   63: 'El compresor Sullair 1 superó la máxima cantidad de horas sin mantenimiento #1', class MTA, trigger "Rec21" bit 13
   64: 'El compresor Sullair 1 superó la máxima cantidad de horas sin mantenimiento #2', class MTA, trigger "Rec21" bit 14
   65: 'El compresor Sullair 1 superó la máxima cantidad de horas sin mantenimiento #3', class MTA, trigger "Rec21" bit 15
   84: 'El compresor Sullair 1 superó la máxima cantidad de horas sin mantenimiento #4', class MTA, trigger "Rec22" bit 8
   85: 'El compresor Sullair 1 superó la máxima cantidad de horas sin mantenimiento #5', class MTA, trigger "Rec22" bit 9
   86: 'El compresor Sullair 0 superó la máxima cantidad de horas sin mantenimiento #1', class MTA, trigger "Rec22" bit 10
   122: 'El compresor Sullair 0 superó la máxima cantidad de horas sin mantenimiento #2', class MTA, trigger "Rec22" bit 11
   123: 'El compresor Sullair 0 superó la máxima cantidad de horas sin mantenimiento #3', class MTA, trigger "Rec22" bit 12
   124: 'El compresor Sullair 0 superó la máxima cantidad de horas sin mantenimiento #4', class MTA, trigger "Rec22" bit 13
   173: 'El compresor Sullair 0 superó la máxima cantidad de horas sin mantenimiento #5', class MTA, trigger "Rec22" bit 14
   174: 'El compresor Atlas 3 superó la máxima cantidad de horas sin mantenimiento #1', class MTA, trigger "Rec22" bit 15
   175: 'El compresor Atlas 3 superó la máxima cantidad de horas sin mantenimiento #2', class MTA, trigger "Rec23" bit 8
   176: 'El compresor Atlas 3 superó la máxima cantidad de horas sin mantenimiento #3', class MTA, trigger "Rec23" bit 9
   177: 'El compresor Atlas 3 superó la máxima cantidad de horas sin mantenimiento #4', class MTA, trigger "Rec23" bit 10
   178: 'El compresor Atlas 3 superó la máxima cantidad de horas sin mantenimiento #5', class MTA, trigger "Rec23" bit 11
   179: 'El compresor Atlas 2 superó la máxima cantidad de horas sin mantenimiento #1', class MTA, trigger "Rec23" bit 12
   180: 'El compresor Atlas 2 superó la máxima cantidad de horas sin mantenimiento #2', class MTA, trigger "Rec23" bit 13
   181: 'El compresor Atlas 2 superó la máxima cantidad de horas sin mantenimiento #3', class MTA, trigger "Rec23" bit 14
   182: 'El compresor Atlas 2 superó la máxima cantidad de horas sin mantenimiento #4', class MTA, trigger "Rec23" bit 15
   183: 'El compresor Atlas 2 superó la máxima cantidad de horas sin mantenimiento #5', class MTA, trigger "Rec24" bit 8
   184: 'El booster 1 superó la máxima cantidad de horas sin mantenimiento', class MTA, trigger "Rec24" bit 9
   185: 'El booster 2 superó la máxima cantidad de horas sin mantenimiento', class MTA, trigger "Rec24" bit 10
   186: 'Temperatura agua de torres compresores elevada', class MTA, trigger "Rec24" bit 11
   187: 'Falla Confirmación de purga - ABC2', class MTA, trigger "Rec17" bit 8
   188: 'Falla Confirmación de purga - ABC3', class MTA, trigger "Rec17" bit 9
   189: 'Falla Confirmación de purga - Bellis', class MTA, trigger "Rec17" bit 10
   190: 'Falla Confirmación de purga - ABC4', class MTA, trigger "Rec17" bit 11
   191: 'Falla Confirmación de purga - ABC5', class MTA, trigger "Rec17" bit 12
   192: 'Falla Confirmación de purga - ABC1', class MTA, trigger "Rec17" bit 13
   199: 'Falla por relé de freq. Comp ALTA', class MTA, trigger "Rec24" bit 15

text list "EstadoMotor": 0 'Detenido'; 1 'En Marcha'; 2 'Arrancando'; 3 'Deteniéndose'; 4 'Espera para Arrancar'; 5 'Sobrecarga de Corriente'; 6 'Deshabilitado'; 7 'En Falla'

text list "EstadoCmpAlta": 256 'Manual'; 512 'Sin Requerimiento'; 1024 'Sin Marcha'; 2048 'En Vacío'; 4096 'En Carga'; 8192 'Manual sin Requerimiento'; 16384 ''; 32768 'Falla'; 1 'Requiere Marcha'

text list "Presostato Ctrl": 0 'Presostato de Control: Desactivado'; 1 'Presostato de Control: Activado'

text list "Presostato de Alarma": 0 'Presostato de Presión Alta: Activado'; 1 'Presostato de Presión Alta: Desactivado'

text list "Lista de rutas": 0 '\Storage Card USB\ABC-1\'; 1 '\Storage Card USB\ABC-2\'; 2 '\Storage Card USB\ABC-3\'; 3 '\Storage Card USB\ABC-4\'; 4 '\Storage Card USB\ABC-5\'; 5 '\Storage Card USB\Bellis\'; 6 '\Storage Card USB\Atlas2\'; 7 '\Storage Card USB\Atlas3\'; 8 '\Storage Card USB\Sullair0\'; 9 '\Storage Card USB\Sullair1\'; 10 '\Storage Card USB\Sullair2\'

text list "Lista de compresores": 0 'ABC-1'; 1 'ABC-2'; 2 'ABC-3'; 3 'ABC-4'; 4 'ABC-5'; 5 'Bellis'; 6 'Atlas 2'; 7 'Atlas 3'; 8 'Sullair 0'; 9 'Sullair 1'; 10 'Sullair 2'

graphic list "Motor2": 0 'Motor2Dorado'; 1 'Motor2Verde_1'; 2 'Motor2VerdeOscuro'; 3 'Motor2Azul'; 4 'Motor2Celeste'; 5 'Motor2Amarillo'; 6 'Motor2Gris_1'; 7 'Motor2Rojo'; 8 'Motor2Dorado'

graphic list "MotorBelliss": 0 'dorado'; 1 'bell1ve'; 2 'bell1ve'; 3 'az'; 4 'az'; 5 'bell1am'; 6 'dorado'; 7 'az'

graphic list "BarraPrioridades": 1 'R1'; 2 'R2'; 3 'R3'; 4 'R4'; 5 'R5'; 6 'R4'; 6 'R6.rlu'

graphic list "Indicador": 0 'indDorado'; 1 'indVerde'; 2 'indVerde_1'; 3 'indAZUL'; 4 'indCeleste'; 5 'indAmarillo'; 6 'indGris'; 7 'indRojo'; 8 'indCeleste'

graphic list "BarraPrioridades_1": 1 'set1'; 2 'set2'; 3 'set3'; 4 'set4'; 5 'set5'; 6 'set4'; 6 'set6'

graphic list "BaseSullChico": 0 'BaseSullChicoDorado_4'; 1 'BaseSullChico'; 2 'BaseSullChico'; 3 'BaseSullChicoAzul_4'; 4 'BaseSullChicoAzul_4'; 5 'BaseSullChicoAmarillo_4'; 6 'BaseSullChicoGris_4'; 7 'BaseSullChicoRojo_4'; 8 'BaseSullChicoAzul_4'

graphic list "MotorTorre": 0 'torreFINAL4C2_1'; 1 'torreFINAL4C2v_2'; 2 'torreFINAL4C2v_2'; 3 'torreFINAL4C2b'; 4 'torreFINAL4C2b'; 5 'torreFINAL4C2a_2'; 6 'torreFINAL4C2_1'; 7 'torreFINAL4C2_1'

graphic list "Secador2": 0 'BaseSullChicoDorado_2'; 1 'BaseSullChico_5'; 2 'BaseSullChico_5'; 3 'BaseSullChicoAzul_2'; 4 'BaseSullChicoAzul_2'; 5 'BaseSullChicoAmarillo_2'; 6 'BaseSullChicoGris_2'; 7 'BaseSullChicoRojo_2'

graphic list "Secador1": 0 'BaseSullChicoDorado_1'; 1 'BaseSullChico_4'; 2 'BaseSullChico_4'; 3 'BaseSullChicoAzul_1'; 4 'BaseSullChicoAzul_1'; 5 'BaseSullChicoAmarillo_1'; 6 'BaseSullChicoGris_1'; 7 'BaseSullChicoRojo_1'

graphic list "Motor Grande": 0 'MotorDorado'; 1 'MotorVerde'; 2 'MotorVerde'; 3 'MotorAzul'; 4 'MotorCeleste'; 5 'MotorAmarillo'; 6 'MotorGris'; 7 'MotorRojo'; 8 'MotorCeleste'

graphic list "Mantenimiento": 0 'MECH2'; 1 'MECH1'

graphic list "Motor Chico": 0 'Booster-D-Dor2'; 1 'Booster-D-VE2'; 2 'Booster-D-VE2'; 3 'Booster-D-Azul2'; 4 'Booster-D-AZ2'; 5 'Booster-D-AM2'; 6 'Booster-D-GR'; 7 'Booster-D-RO2'; 8 'Booster-D-AZ2'

graphic list "Hélice": 0 'Booster-C1'; 1 'Booster-C2'

screen "Graf-Corrientes" 1280x800, template "Plantilla"
   TrendView "Visor de curvas_1" at 8,72 size 1260x636
   TextField "Campo de texto_16" at 493,10 size 294x27; Text 'Gráficas - Sentron Pac - Corrientes'

screen "Graf-Fase" 1280x800, template "Plantilla"
   TrendView "Visor de curvas_1" at 3,65 size 1268x644
   TextField "Campo de texto_16" at 477,10 size 364x27; Text 'Gráficas - Sentron Pac - Tensiones de Fase'

screen "Grafica" 1280x800, template "Plantilla"
   Button "Botón_7" at 368,280 size 240x49; TextOff 'Presión Baja'
      on Click: ActivateScreen("GraficaPBAJA", 0)
   Button "Botón_12" at 367,440 size 240x49; TextOff 'Temperatura Chillers'
      on Click: ActivateScreen("GraficaTCH", 0)
   Button "Botón_13" at 368,216 size 240x49; TextOff 'Presión Alta'
      on Click: ActivateScreen("GraficaPALTA", 0)
   TextField "Campo de texto_1" at 55,108 size 353x27; Text 'Seleccione la variable que desea graficar:'
   Button "Botón_1" at 767,280 size 240x49; TextOff 'Todas Cavaleto'
      on Click: ActivateScreen("GraficaTodas", 0)
   TextField "Campo de texto_16" at 521,10 size 226x27; Text 'Graficar variable analógica'
   Button "Botón_2" at 368,344 size 240x49; TextOff 'Temperatura Cavaleto'
      on Click: ActivateScreen("GraficaTCAV", 0)
   Button "Botón_3" at 766,440 size 240x49; TextOff 'Grafico Caudal/Potencia'
      on Click: ActivateScreen("Graf-cau-pot-actual", 0)
   Button "Botón_4" at 769,526 size 240x49; TextOff 'Historico Caudal/Potencia'
      on Click: ActivateScreen("Graf-cau-pot-historico", 0)

screen "GraficaPALTA" 1280x800, template "Plantilla"
   TrendView "Visor de curvas_1" at 5,79 size 1234x618
   TextField "Campo de texto_16" at 521,10 size 193x27; Text 'Grafica Presión de Alta'

screen "GraficaPBAJA" 1280x800, template "Plantilla"
   TrendView "Visor de curvas_1" at 5,71 size 1242x626
   TextField "Campo de texto_16" at 521,10 size 198x27; Text 'Grafica Presión de Baja'

screen "GraficaTCAV" 1280x800, template "Plantilla"
   TrendView "Visor de curvas_1" at 5,71 size 1242x626
   TextField "Campo de texto_16" at 521,10 size 254x27; Text 'Grafica Temperatura Cavaleto'

screen "GraficaTCH" 1280x800, template "Plantilla"
   TrendView "Visor de curvas_1" at 5,71 size 1242x626
   TextField "Campo de texto_16" at 521,10 size 243x27; Text 'Grafica Temperatura Chillers'

screen "GraficaTodas" 1280x800, template "Plantilla"
   TrendView "Visor de curvas_1" at 5,71 size 1242x626

screen "Graf-Linea" 1280x800, template "Plantilla"
   TrendView "Visor de curvas_1" at 3,65 size 1268x652
   TextField "Campo de texto_16" at 453,10 size 370x27; Text 'Gráficas - Sentron Pac - Tensiones de Línea'

screen "Graf-Pot" 1280x800, template "Plantilla"
   TrendView "Visor de curvas_1" at 3,65 size 1268x644
   TextField "Campo de texto_16" at 477,10 size 339x27; Text 'Gráficas - Sentron Pac - Potencia x Fase'

screen "Graf-PotTotal" 1280x800, template "Plantilla"
   TrendView "Visor de curvas_1" at 3,65 size 1268x644
   TextField "Campo de texto_16" at 477,10 size 327x27; Text 'Gráficas - Sentron Pac - Potencia Total'

screen "IluminaciónMTA" 1280x800, template "Plantilla"
   Polygon "Polígono_6" at 1018,121 size 183x209
      Visibility <- "ON"
   Ellipse "Elipse_4" at 1019,317 size 184x29
      Visibility <- "ON"
   Polygon "Polígono_3" at 782,137 size 351x377
      Visibility <- "ON"
   Ellipse "Elipse_5" at 789,485 size 344x61
      Visibility <- "ON"
   Polygon "Polígono_2" at 446,161 size 559x577
      Visibility <- "ON"
   Ellipse "Elipse_1" at 694,118 size 59x74
      Appearance <- "ON"
   Ellipse "Elipse_2" at 940,112 size 35x50
      Appearance <- "ON"
   Ellipse "Elipse_3" at 1100,112 size 19x26
      Appearance <- "ON"
   Switch "Interruptor_1" at 36,546 size 510x96; TextOff 'Encendido Permanente OFF'; CaptionText 'Switch'; TextOn 'Encendido Permanente ON'
      Appearance <- "MantenerON"
      ProcessValue <- "MantenerON"
   Button "Botón_1" at 36,264 size 248x96; TextOff 'Encender'
      on Press: SetBit("EncendidoPanel")
      on Release: ResetBit("EncendidoPanel")
   Button "Botón_2" at 298,263 size 248x96; TextOff 'Apagar'
      on Press: SetBit("ApagadoPanel")
      on Release: ResetBit("ApagadoPanel")
   IOField "Campo ES_1" at 257,148 size 140x39; FormatPattern 99; Unit    Min.
      ProcessValue <- "TiempoIluminación"
   TextField "Campo de texto_1" at 42,156 size 186x27; Text 'Tiempo de encendido'
   TextField "Campo de texto_3" at 58,190 size 466x58; Text 'La iluminación puede ser encendida desde el panel o desde el pulsador. En caso de no ser apagada mediante los mismos medios, el PLC la apagará automáticamente al concluir el "tiempo de encendido".'
   TextField "Campo de texto_2" at 58,414 size 433x112; Text 'En caso de necesitar permanecer con la iluminación encendida durante un tiempo mayor al "tiempo de encendido", se provee la posibilidad de seleccionar el "encendido permanente". Mientras el "encendido permanente" esté activado la iluminación se mantendrá encendida, y el PLC dejará de controlar el apagado automático.'
   TextField "Campo de texto_16" at 553,10 size 177x27; Text 'Iluminación Cavaleto'

screen "INICIO" 1280x800, template "Plantilla"
   Button "Botón_1" at 1025,513 size 108x65; TextOff 'Cerrar Runtime'; Authorization "Administración de usuarios"
      on Press: StopRuntime(0)
   Button "Botón_2" at 115,501 size 130x47; TextOff 'Iniciar Sesion'; PictureOff "Gráfico_5"
      on Click: function_a2a04561()
   UserView "Visor de usuarios_1" at 266,510 size 665x23
   GraphicView "Visor de gráficos_1" at 96,110 size 1064x352; Picture "banner-home"
   Button "Botón_3" at 115,557 size 130x47; TextOff 'Cerrar Sesion'; PictureOff "Gráfico_5"
      on Click: function_f23ef4c9()
   Button "Botón_4" at 802,557 size 130x47; TextOff 'Administrar'; Authorization "Administración de usuarios"; PictureOff "Gráfico_5"
      on Click: ActivateScreen("INICIO-Administración", 0)

screen "INICIO-Administración" 1280x800, template "Plantilla"
   Button "Botón_1" at 1025,513 size 108x65; TextOff 'Cerrar Runtime'; Authorization "Administración de usuarios"
      on Press: StopRuntime(0)
   Button "Botón_2" at 115,501 size 130x47; TextOff 'Iniciar Sesion'; PictureOff "Gráfico_5"
      on Click: function_a2a04561()
   UserView "Visor de usuarios_1" at 266,502 size 665x23
   GraphicView "Visor de gráficos_1" at 96,110 size 1064x352; Picture "banner-home"
   Button "Botón_3" at 115,557 size 130x47; TextOff 'Cerrar Sesion'; PictureOff "Gráfico_5"
      on Click: function_f23ef4c9()
   UserView "Visor de usuarios_2" at 266,534 size 665x143

screen "MTA-ALTAMC001" 1280x800, template "Plantilla-Alta-Cmp"
   Switch "Interruptor_1" at 156,166 size 37x37; TextOn '1'; TextOff '0'; CaptionText 'Switch'; PictureOff "A2"; Authorization "Operación"; PictureOn "A"
      ProcessValue <- "Auto1"
      Visibility <- "MantMC001"
   Button "Botón_6" at 27,153 size 88x62; TextOff 'ABC 2'
   ScreenModuleView "Faceplate_6_1" at 348,235 size 76x34; ScreenModuleType ""
      Guid_{11997190-52606} <- "IndV1"
      Guid_{11997190-52610} <- "IndR1"
      Guid_{11997190-52608} <- "IndVparp1"
   ScreenModuleView "Faceplate_7_1" at 208,157 size 216x70
      Guid_{11997190-23983} <- "ParadaMC001"
      Guid_{11997190-23981} <- "MarchaMC001"
      Guid_{11997190-90329} <- "ForzarParada1"
      Guid_{11997190-180841} <- "MantMC001"
      Guid_{11997190-89807} <- "SPOFFF1"
      Guid_{11997190-89795} <- "ForzandoMarcha1"
      Guid_{11997190-90325} <- "MarchaMC001"
      Guid_{11997190-88662} <- "MarchaOK1"
      Guid_{11997190-23985} <- "AnimMenuMC001"
      Guid_{11997190-89805} <- "SPONF1"
   GraphicIOField "Campo ES gráfico_2" at 16,279 size 422x6; PictureList "Indicador"
      ProcessValue <- "AnimMotorMC001"
   SymbolicIOField "Campo ES simbólico_4" at 25,245 size 290x21; TextOff '0'; TextOn '1'; TextList "EstadoMotor"
      ProcessValue <- "AnimMotorMC001"
   TextField "Campo de texto_1" at 272,362 size 72x27; Text 'Seteada'
   Button "Botón_1" at 192,442 size 48x38; TextOff 'Incrementar'; Authorization "Operación"; PictureOff "Gráfico_3"
      on Press: SetBit("IncP1")
      on Release: ResetBit("IncP1")
   Button "Botón_2" at 192,402 size 48x38; TextOff 'Decrementar'; Authorization "Operación"; PictureOff "Gráfico_1"
      on Press: SetBit("DecP1")
      on Release: ResetBit("DecP1")
   TextField "Campo de texto_2" at 88,426 size 84x27; Text 'Prioridad'
   GraphicIOField "Campo ES gráfico_1" at 300,402 size 16x78; PictureList "BarraPrioridades"
      ProcessValue <- "VCMP1"
   GraphicIOField "Campo ES gráfico_4" at 380,402 size 16x78; PictureList "BarraPrioridades_1"
      ProcessValue <- "PriRealCMP1"
   TextField "Campo de texto_10" at 368,363 size 40x27; Text 'Real'
   SymbolicIOField "Campo ES simbólico_1" at 15,290 size 424x37; TextOff '0'; TextOn '1'; TextList "EstadoCmpAlta"
      ProcessValue <- "Est1"
      Visibility <- "MantMC001"
   Button "Botón_3" at 396,106 size 40x38; TextOff 'Text'; PictureOff "x"
      on Click: function_efd93a16()
   Button "Botón_4" at 306,600 size 96x35; TextOff 'Hecho'; Authorization "Administración de usuarios"
      on Press: SetTag("Varios_UltimoMantMC001_1", "HORAS1")
   TextField "Campo de texto_6" at 32,510 size 326x27; Text 'Tiempo de funcionamiento acumulado'
   TextField "Campo de texto_3" at 32,343 size 158x27; Text 'Seteo de Prioridad'
   TextField "Campo de texto_16" at 521,10 size 279x27; Text 'Menú Compresor ABC-2 (MC001)'
   Button "Botón_5" at 306,665 size 96x35; TextOff 'Hecho'; Authorization "Administración de usuarios"
      on Press: SetTag("Varios_UltimoMantMC001_2", "HORAS1")
   TextField "Campo de texto_4" at 32,570 size 231x27; Text 'Próximo mantenimiento #1'
   TextField "Campo de texto_5" at 32,635 size 231x27; Text 'Próximo mantenimiento #2'
   Switch "Interruptor_2" at 459,548 size 120x40; TextOff 'OFF'; TextOn 'ON'; CaptionText 'Switch'
      ProcessValue <- "DB-PurgaComAlta_Habil_PurgaABC2"
   IOField "Campo ES_4" at 574,609 size 96x32; FormatPattern 99; Unit  min
      ProcessValue <- "DB-PurgaComAlta_Toff_PurgaABC2"
   IOField "Campo ES_5" at 574,654 size 96x32; FormatPattern 99; Unit  seg
      ProcessValue <- "DB-PurgaComAlta_Ton_PurgaABC2"
   TextField "Campo de texto_7" at 459,613 size 97x27; Text 'Tiempo Off'
   TextField "Campo de texto_8" at 459,655 size 96x27; Text 'Tiempo On'
   Button "Botón_7" at 595,548 size 80x40; TextOff 'Prueba'
      on Press: SetBit("DB-PurgaComAlta_Prueba_PurgaABC2")
      on Release: ResetBit("DB-PurgaComAlta_Prueba_PurgaABC2")
      Appearance <- "MC001_EVP"
      ObjectEnable <- "MC001_EVP"
   TextField "Campo de texto_9" at 456,510 size 131x27; Text 'Ciclo de Purga:'
   IOField "Campo ES_7" at 20,535 size 173x35; Authorization "Administración de usuarios"; FormatPattern 999999999; Unit  hs
      ProcessValue <- "HORAS1"
      Appearance <- "EstadoMantMC001"
   IOField "Campo ES_1" at 200,535 size 80x35; Authorization "Administración de usuarios"; FormatPattern 99; Unit  min
      ProcessValue <- "MIN1"
   IOField "Campo ES_2" at 20,595 size 173x35; FormatPattern 999999999; Unit  hs
      ProcessValue <- "ProxMantMC001_1"
      Appearance <- "LimiteMantMC001_1"
   IOField "Campo ES_3" at 20,660 size 173x35; FormatPattern 999999999; Unit  hs
      ProcessValue <- "ProxMantMC001_2"
      Appearance <- "LimiteMantMC001_2"

screen "MTA-ALTAMC002" 1280x800, template "Plantilla-Alta-Cmp"
   TextField "Campo de texto_1" at 266,362 size 72x27; Text 'Seteada'
   TextField "Campo de texto_2" at 82,426 size 84x27; Text 'Prioridad'
   TextField "Campo de texto_10" at 362,363 size 40x27; Text 'Real'
   TextField "Campo de texto_6" at 32,510 size 326x27; Text 'Tiempo de funcionamiento acumulado'
   TextField "Campo de texto_3" at 26,343 size 158x27; Text 'Seteo de Prioridad'
   Button "Botón_1" at 186,442 size 48x38; TextOff 'Incrementar'; Authorization "Operación"; PictureOff "Gráfico_3"
      on Press: SetBit("IncP2")
      on Release: ResetBit("IncP2")
   Button "Botón_2" at 186,402 size 48x38; TextOff 'Decrementar'; Authorization "Operación"; PictureOff "Gráfico_1"
      on Press: SetBit("DecP2")
      on Release: ResetBit("DecP2")
   Button "Botón_3" at 390,106 size 40x38; TextOff 'Text'; PictureOff "x"
      on Click: function_efd93a16()
   Button "Botón_4" at 306,600 size 96x35; TextOff 'Hecho'; Authorization "Administración de usuarios"
      on Press: SetTag("Varios_UltimoMantMC002_1", "HORAS2")
   GraphicIOField "Campo ES gráfico_1" at 294,402 size 16x78; PictureList "BarraPrioridades"
      ProcessValue <- "VCMP2"
   GraphicIOField "Campo ES gráfico_4" at 374,402 size 16x78; PictureList "BarraPrioridades_1"
      ProcessValue <- "PriRealCMP2"
   SymbolicIOField "Campo ES simbólico_1" at 9,290 size 424x37; TextOff '0'; TextOn '1'; TextList "EstadoCmpAlta"
      ProcessValue <- "Est2"
      Visibility <- "MantMC002"
   TextField "Campo de texto_16" at 521,10 size 279x27; Text 'Menú Compresor ABC-3 (MC002)'
   TextField "Campo de texto_4" at 32,570 size 231x27; Text 'Próximo mantenimiento #1'
   TextField "Campo de texto_5" at 32,635 size 231x27; Text 'Próximo mantenimiento #2'
   Button "Botón_5" at 306,665 size 96x35; TextOff 'Hecho'; Authorization "Administración de usuarios"
      on Press: SetTag("Varios_UltimoMantMC002_2", "HORAS2")
   IOField "Campo ES_4" at 574,609 size 96x32; FormatPattern 99; Unit  min
      ProcessValue <- "DB-PurgaComAlta_Toff_PurgaABC3"
   IOField "Campo ES_5" at 574,654 size 96x32; FormatPattern 99; Unit  seg
      ProcessValue <- "DB-PurgaComAlta_Ton_PurgaABC3"
   TextField "Campo de texto_7" at 459,613 size 97x27; Text 'Tiempo Off'
   TextField "Campo de texto_8" at 459,655 size 96x27; Text 'Tiempo On'
   Switch "Interruptor_2" at 459,548 size 120x40; TextOff 'OFF'; CaptionText 'Switch'; TextOn 'ON'
      ProcessValue <- "DB-PurgaComAlta_Habil_PurgaABC3"
   Button "Botón_7" at 595,548 size 80x40; TextOff 'Prueba'
      on Press: SetBit("DB-PurgaComAlta_Prueba_PurgaABC3")
      on Release: ResetBit("DB-PurgaComAlta_Prueba_PurgaABC3")
      Appearance <- "MC002_EVP"
      ObjectEnable <- "MC002_EVP"
   TextField "Campo de texto_9" at 456,510 size 131x27; Text 'Ciclo de Purga:'
   GraphicIOField "Campo ES gráfico_2" at 10,279 size 422x6; PictureList "Indicador"
      ProcessValue <- "AnimMotorMC002"
   SymbolicIOField "Campo ES simbólico_4" at 19,245 size 290x21; TextOff '0'; TextOn '1'; TextList "EstadoMotor"
      ProcessValue <- "AnimMotorMC002"
   Button "Botón_6" at 21,153 size 88x62; TextOff 'ABC 3'
   Switch "Interruptor_1" at 150,166 size 37x37; TextOn '1'; TextOff '0'; CaptionText 'Switch'; PictureOff "A2"; Authorization "Operación"; PictureOn "A"
      ProcessValue <- "Auto2"
      Visibility <- "MantMC002"
   ScreenModuleView "Faceplate_6_1" at 342,235 size 76x34; ScreenModuleType ""
      Guid_{11997190-52606} <- "IndV2"
      Guid_{11997190-52610} <- "IndR2"
      Guid_{11997190-52608} <- "IndVparp2"
   ScreenModuleView "Faceplate_7_1" at 212,161 size 208x70
      Guid_{11997190-23983} <- "ParadaMC002"
      Guid_{11997190-23981} <- "MarchaMC002"
      Guid_{11997190-90329} <- "ForzarParada2"
      Guid_{11997190-180841} <- "MantMC002"
      Guid_{11997190-89807} <- "SPOFFF2"
      Guid_{11997190-89795} <- "ForzandoMarcha2"
      Guid_{11997190-90325} <- "MarchaMC002"
      Guid_{11997190-88662} <- "MarchaOK2"
      Guid_{11997190-23985} <- "AnimMenuMC002"
      Guid_{11997190-89805} <- "SPONF2"
   IOField "Campo ES_7" at 20,535 size 173x35; Authorization "Administración de usuarios"; FormatPattern 999999999; Unit  hs
      ProcessValue <- "HORAS2"
      Appearance <- "EstadoMantMC002"
   IOField "Campo ES_1" at 200,535 size 80x35; Authorization "Administración de usuarios"; FormatPattern 99; Unit  min
      ProcessValue <- "MIN2"
   IOField "Campo ES_2" at 20,595 size 173x35; FormatPattern 999999999; Unit  hs
      ProcessValue <- "ProxMantMC002_1"
      Appearance <- "LimiteMantMC002_1"
   IOField "Campo ES_3" at 20,660 size 173x35; FormatPattern 999999999; Unit  hs
      ProcessValue <- "ProxMantMC002_2"
      Appearance <- "LimiteMantMC002_2"

screen "MTA-ALTAMC003" 1280x800, template "Plantilla-Alta-Cmp"
   Switch "Interruptor_1" at 150,119 size 37x37; TextOn '1'; TextOff '0'; CaptionText 'Switch'; PictureOff "A2"; Authorization "Operación"; PictureOn "A"
      ProcessValue <- "Auto3"
      Visibility <- "MantMC003"
   Button "Botón_6" at 13,106 size 88x62; TextOff 'Bellis'
   ScreenModuleView "Faceplate_6_1" at 342,236 size 76x34; ScreenModuleType ""
      Guid_{11997190-52606} <- "IndV3"
      Guid_{11997190-52610} <- "IndR3"
      Guid_{11997190-52608} <- "IndVparp3"
   Button "Botón_1" at 186,441 size 48x38; TextOff 'Incrementar'; Authorization "Operación"; PictureOff "Gráfico_3"
      on Press: SetBit("IncP3")
      on Release: ResetBit("IncP3")
   Button "Botón_2" at 186,401 size 48x38; TextOff 'Decrementar'; Authorization "Operación"; PictureOff "Gráfico_1"
      on Press: SetBit("DecP3")
      on Release: ResetBit("DecP3")
   TextField "Campo de texto_6" at 266,362 size 72x27; Text 'Seteada'
   TextField "Campo de texto_7" at 82,426 size 84x27; Text 'Prioridad'
   TextField "Campo de texto_8" at 362,363 size 40x27; Text 'Real'
   TextField "Campo de texto_9" at 32,510 size 326x27; Text 'Tiempo de funcionamiento acumulado'
   TextField "Campo de texto_11" at 26,343 size 158x27; Text 'Seteo de Prioridad'
   Button "Botón_7" at 390,58 size 40x38; TextOff 'Text'; PictureOff "x"
      on Click: function_efd93a16()
   Button "Botón_8" at 306,600 size 96x35; TextOff 'Hecho'; Authorization "Administración de usuarios"
      on Press: SetTag("Varios_UltimoMantMC003_1", "HORAS3")
   GraphicIOField "Campo ES gráfico_3" at 294,402 size 16x78; PictureList "BarraPrioridades"
      ProcessValue <- "VCMP3"
   GraphicIOField "Campo ES gráfico_5" at 374,402 size 16x78; PictureList "BarraPrioridades_1"
      ProcessValue <- "PriRealCMP3"
   SymbolicIOField "Campo ES simbólico_2" at 9,290 size 424x37; TextOff '0'; TextOn '1'; TextList "EstadoCmpAlta"
      ProcessValue <- "Est3"
      Visibility <- "MantMC003"
   TextField "Campo de texto_16" at 521,10 size 270x27; Text 'Menú Compresor Bellis (MC003)'
   IOField "Campo ES_2" at 606,443 size 88x23; FormatPattern 99; Unit  Min.
      ProcessValue <- "TiempoMaxBellismedia"
   TextField "Campo de texto_1" at 447,428 size 143x50; Text 'Tiempo máximo en Media Carga'
   Button "Botón_3" at 306,665 size 96x35; TextOff 'Hecho'; Authorization "Administración de usuarios"
      on Press: SetTag("Varios_UltimoMantMC003_2", "HORAS3")
   TextField "Campo de texto_4" at 32,570 size 231x27; Text 'Próximo mantenimiento #1'
   TextField "Campo de texto_5" at 32,635 size 231x27; Text 'Próximo mantenimiento #2'
   IOField "Campo ES_5" at 574,609 size 96x32; FormatPattern 99; Unit  min
      ProcessValue <- "DB-PurgaComAlta_Toff_PurgaBallis"
   IOField "Campo ES_6" at 574,654 size 96x32; FormatPattern 99; Unit  seg
      ProcessValue <- "DB-PurgaComAlta_Ton_PurgaBallis"
   TextField "Campo de texto_2" at 459,613 size 97x27; Text 'Tiempo Off'
   TextField "Campo de texto_3" at 459,655 size 96x27; Text 'Tiempo On'
   Switch "Interruptor_3" at 459,548 size 120x40; TextOff 'OFF'; CaptionText 'Switch'; TextOn 'ON'
      ProcessValue <- "DB-PurgaComAlta_Habil_PurgaBallis"
   Button "Botón_4" at 595,548 size 80x40; TextOff 'Prueba'
      on Press: SetBit("DB-PurgaComAlta_Prueba_PurgaBallis")
      on Release: ResetBit("DB-PurgaComAlta_Prueba_PurgaBallis")
      ObjectEnable <- "MC003_EVP"
      Appearance <- "MC003_EVP"
   TextField "Campo de texto_10" at 456,510 size 131x27; Text 'Ciclo de Purga:'
   GraphicIOField "Campo ES gráfico_2" at 10,280 size 422x6; PictureList "Indicador"
      ProcessValue <- "AnimMotorMC003"
   SymbolicIOField "Campo ES simbólico_4" at 19,246 size 290x21; TextOff '0'; TextOn '1'; TextList "EstadoMotor"
      ProcessValue <- "AnimMotorMC003"
   IOField "Campo ES_7" at 20,535 size 173x35; Authorization "Administración de usuarios"; FormatPattern 999999999; Unit  hs
      ProcessValue <- "HORAS3"
      Appearance <- "EstadoMantMC003"
   IOField "Campo ES_1" at 200,535 size 80x35; Authorization "Administración de usuarios"; FormatPattern 99; Unit  min
      ProcessValue <- "MIN3"
   IOField "Campo ES_3" at 20,595 size 173x35; FormatPattern 999999999; Unit  hs
      ProcessValue <- "ProxMantMC003_1"
      Appearance <- "LimiteMantMC003_1"
   IOField "Campo ES_4" at 20,660 size 173x35; FormatPattern 999999999; Unit  hs
      ProcessValue <- "ProxMantMC003_2"
      Appearance <- "LimiteMantMC003_2"
   Switch "Interruptor_2" at 19,168 size 160x36; TextOn 'Media Carga'; TextOff 'Carga Completa'; CaptionText 'Switch'; Authorization "Operación"
      ProcessValue <- "MediaCargaBellis"
   ScreenModuleView "Faceplate_10_1" at 206,110 size 209x118
      Guid_{11997190-23983} <- "ParadaMC003"
      Guid_{11997190-88662} <- "MarchaOK3"
      Guid_{11997190-23981} <- "MarchaMC003"
      Guid_{11997190-90329} <- "ForzarParada3"
      Guid_{11997190-116346} <- "SPOFFF3b"
      Guid_{11997190-89807} <- "SPOFFF3"
      Guid_{11997190-89795} <- "ForzandoMarcha3"
      Guid_{11997190-90325} <- "MarchaMC003"
      Guid_{11997190-116342} <- "SPONF3b"
      Guid_{11997190-23985} <- "AnimMenuMC003"
      Guid_{11997190-89805} <- "SPONF3"

screen "MTA-ALTAMC004" 1280x800, template "Plantilla-Alta-Cmp"
   Button "Botón_1" at 186,441 size 48x38; TextOff 'Incrementar'; Authorization "Operación"; PictureOff "Gráfico_3"
      on Press: SetBit("IncP4")
      on Release: ResetBit("IncP4")
   Button "Botón_2" at 186,401 size 48x38; TextOff 'Decrementar'; Authorization "Operación"; PictureOff "Gráfico_1"
      on Press: SetBit("DecP4")
      on Release: ResetBit("DecP4")
   Button "Botón_7" at 390,106 size 40x38; TextOff 'Text'; PictureOff "x"
      on Click: function_efd93a16()
   Button "Botón_8" at 300,600 size 96x35; TextOff 'Hecho'; Authorization "Administración de usuarios"
      on Press: SetTag("Varios_UltimoMantMC004_1", "HORAS4")
   TextField "Campo de texto_6" at 266,362 size 72x27; Text 'Seteada'
   TextField "Campo de texto_7" at 82,426 size 84x27; Text 'Prioridad'
   TextField "Campo de texto_8" at 362,363 size 40x27; Text 'Real'
   TextField "Campo de texto_11" at 26,343 size 158x27; Text 'Seteo de Prioridad'
   GraphicIOField "Campo ES gráfico_3" at 294,402 size 16x78; PictureList "BarraPrioridades"
      ProcessValue <- "VCMP4"
   GraphicIOField "Campo ES gráfico_5" at 374,402 size 16x78; PictureList "BarraPrioridades_1"
      ProcessValue <- "PriRealCMP4"
   SymbolicIOField "Campo ES simbólico_2" at 9,290 size 424x37; TextOff '0'; TextOn '1'; TextList "EstadoCmpAlta"
      ProcessValue <- "Est4"
      Visibility <- "MantMC004"
   TextField "Campo de texto_16" at 521,10 size 279x27; Text 'Menú Compresor ABC-4 (MC004)'
   TextField "Campo de texto_1" at 32,510 size 326x27; Text 'Tiempo de funcionamiento acumulado'
   TextField "Campo de texto_4" at 32,570 size 231x27; Text 'Próximo mantenimiento #1'
   TextField "Campo de texto_5" at 32,635 size 231x27; Text 'Próximo mantenimiento #2'
   Button "Botón_3" at 300,665 size 96x35; TextOff 'Hecho'; Authorization "Administración de usuarios"
      on Press: SetTag("Varios_UltimoMantMC004_2", "HORAS4")
   IOField "Campo ES_4" at 574,609 size 96x32; FormatPattern 99; Unit  min
      ProcessValue <- "DB-PurgaComAlta_Toff_PurgaABC4"
   IOField "Campo ES_5" at 574,654 size 96x32; FormatPattern 99; Unit  seg
      ProcessValue <- "DB-PurgaComAlta_Ton_PurgaABC4"
   TextField "Campo de texto_2" at 459,613 size 97x27; Text 'Tiempo Off'
   TextField "Campo de texto_3" at 459,655 size 96x27; Text 'Tiempo On'
   Switch "Interruptor_2" at 459,548 size 120x40; TextOff 'OFF'; TextOn 'ON'; CaptionText 'Switch'
      ProcessValue <- "DB-PurgaComAlta_Habil_PurgaABC4"
   Button "Botón_4" at 595,548 size 80x40; TextOff 'Prueba'
      on Press: SetBit("DB-PurgaComAlta_Prueba_PurgaABC4")
      on Release: ResetBit("DB-PurgaComAlta_Prueba_PurgaABC4")
      ObjectEnable <- "MC004_EVP"
      Appearance <- "MC004_EVP"
   TextField "Campo de texto_9" at 456,510 size 131x27; Text 'Ciclo de Purga:'
   GraphicIOField "Campo ES gráfico_2" at 10,280 size 422x6; PictureList "Indicador"
      ProcessValue <- "AnimMotorMC004"
   SymbolicIOField "Campo ES simbólico_4" at 19,246 size 290x21; TextOff '0'; TextOn '1'; TextList "EstadoMotor"
      ProcessValue <- "AnimMotorMC004"
   Button "Botón_6" at 13,154 size 88x62; TextOff 'ABC 4'
   Switch "Interruptor_1" at 150,167 size 37x37; TextOn '1'; TextOff '0'; CaptionText 'Switch'; PictureOff "A2"; Authorization "Operación"; PictureOn "A"
      ProcessValue <- "Auto4"
      Visibility <- "MantMC004"
   ScreenModuleView "Faceplate_6_1" at 342,236 size 76x34; ScreenModuleType ""
      Guid_{11997190-52606} <- "IndV4"
      Guid_{11997190-52610} <- "IndR4"
      Guid_{11997190-52608} <- "IndVparp4"
   ScreenModuleView "Faceplate_7_1" at 213,158 size 208x70
      Guid_{11997190-23983} <- "ParadaMC004"
      Guid_{11997190-23981} <- "MarchaMC004"
      Guid_{11997190-90329} <- "ForzarParada4"
      Guid_{11997190-180841} <- "MantMC004"
      Guid_{11997190-89807} <- "SPOFFF4"
      Guid_{11997190-89795} <- "ForzandoMarcha4"
      Guid_{11997190-90325} <- "MarchaMC004"
      Guid_{11997190-88662} <- "MarchaOK4"
      Guid_{11997190-23985} <- "AnimMenuMC004"
      Guid_{11997190-89805} <- "SPONF4"
   IOField "Campo ES_7" at 20,535 size 173x35; Authorization "Administración de usuarios"; FormatPattern 999999999; Unit  hs
      ProcessValue <- "HORAS4"
      Appearance <- "EstadoMantMC004"
   IOField "Campo ES_1" at 200,535 size 80x35; Authorization "Administración de usuarios"; FormatPattern 99; Unit  min
      ProcessValue <- "MIN4"
   IOField "Campo ES_2" at 20,595 size 173x35; FormatPattern 999999999; Unit  hs
      ProcessValue <- "ProxMantMC004_1"
      Appearance <- "LimiteMantMC004_1"
   IOField "Campo ES_3" at 20,660 size 173x35; FormatPattern 999999999; Unit  hs
      ProcessValue <- "ProxMantMC004_2"
      Appearance <- "LimiteMantMC004_2"

